(* Logix 5000 project; controller PLC_MCC1300_75F1 vendor 1 type 14 code 166 rev 32.11; software revision 32.04; part 77 of 83 *)
(* tags used below, declared in another part *)
   CM_AreaStackerToLine_JS1_Sync : CM_AreaStackerToLine;
   CM_ConveyorStackerToLine_JS1_Sync : CM_ConveyorStackerToLine;
   CONST_tPlant : UDT_PLANT_CONSTANTS;
   GP_AccessArea_M311S : GP_AccessArea;
   GP_AccessArea_M311S_STC : GP_AccessArea_STC;
   GP_AccessArea_M316S : GP_AccessArea;
   GP_AccessArea_M316S_STC : GP_AccessArea_STC;
   GP_OB_InitializeMain : GP_OB_Initialize;
   GP_TrackingGetLength : GP_TrackingGetLength;
   M302SpeedUp : MAC_SpeedUp;
   M30xTrimDeck : MAC_TrimmingDeck[5];
   M310B : MAC_Conveyor;
   M310B_ALM : MAC_Conveyor_ALM;
   M310B_HMW : MAC_Conveyor_HMW;
   M310Popup : MAC_Popup_ZC[2];
   M311 : MAC_Conveyor;
   M311_ALM : MAC_Conveyor_ALM;
   M311_HMW : MAC_Conveyor_HMW;
   M311A : MAC_Rotator;
   M311A_ALM : MAC_Rotator_ALM;
   M312 : MAC_Conveyor_Single;
   M312_ALM : MAC_Conveyor_ALM;
   M312_HMW : MAC_Conveyor_HMW;
   M316 : MAC_Conveyor;
   M316A : MAC_Rotator;
   M317 : MAC_Conveyor_Single;
   xAlwaysON : BOOL;
   Z300_Conveyor : UDT_StandConv[29];
   Z300_Conveyor_ALM : MAC_Conveyor_ZC_ALM[29];
   Z300_Conveyor_HMW : MAC_Conveyor_ZC_HMW[29];
   Z300_LineTracking : UDT_LINE_TRACKING;
   Z301 : MAC_Zone_ML;
   Z301_HMR : MAC_Zone_ML_HMR;
   Z301_HMW : MAC_Zone_ML_HMW;
   Z311S : MAC_SafetyAccess;
   Z311S_ALM : MAC_SafetyAccess_ALM;
   Z311S_HMR : MAC_SafetyAccess_HMR;
   Z311S_INPUT_xAccessReqRotator : BOOL;
   Z311S_INPUT_xSafetyAreaRotator : BOOL;
   Z311S_OUTPUT_xEL_AccessAcceptedRotator : BOOL;
   Z311S_OUTPUT_xHL_AccessAcceptedRotator : BOOL;
   Z311S_OUTPUT_xHL_SafetyAreaRotatorNOK : BOOL;
   Z316S : MAC_SafetyAccess;
   Z316S_ALM : MAC_SafetyAccess_ALM;
   Z316S_HMR : MAC_SafetyAccess_HMR;
   Z316S_INPUT_xAccessReqRotator : BOOL;
   Z316S_INPUT_xSafetyAreaRotator : BOOL;
   Z316S_OUTPUT_xEL_AccessAcceptedRotator : BOOL;
   Z316S_OUTPUT_xHL_AccessAcceptedRotator : BOOL;
   Z316S_OUTPUT_xHL_SafetyAreaRotatorNOK : BOOL;
   Z401 : MAC_Zone;
   Z401_ALM : MAC_Zone_ALM;
   Z401_HMR : MAC_Zone_HMR;
   Z401_HMW : MAC_Zone_HMW;
   Z401_INPUT_xMainLineEmergencyON : BOOL;
   Z401_OUTPUT_xMCC_SafetyPanel1 : BOOL;
   Z402 : MAC_Zone;
(* MainProgram, continued *)

   54: XIC(Z300_Conveyor_HMW[7].xLocalCleaningRequest)XIC(Z300_Conveyor[0].tIN_Zone.xCleanZoneAccepted)OTE(Z300_Conveyor_HMW[8].xLocalCleaningRequest);
   // M312 Cleaning Enabled
   55: XIC(Z300_Conveyor_HMW[8].xLocalCleaningRequest)XIC(Z300_Conveyor[0].tIN_Zone.xCleanZoneAccepted)[OTE(Z300_Conveyor_HMW[9].xLocalCleaningRequest) ,OTE(Z300_Conveyor_HMW[10].xLocalCleaningRequest) ];
   56: XIC(Z300_Conveyor_HMW[10].xLocalCleaningRequest)XIC(Z300_Conveyor[0].tIN_Zone.xCleanZoneAccepted)OTE(Z300_Conveyor_HMW[11].xLocalCleaningRequest);
   57: XIC(Z301.ST_xReqCleaning)XIC(Z300_Conveyor[0].ST_xCleaningConditionOK)XIC(Z300_Conveyor[1].ST_xCleaningConditionOK)XIC(Z300_Conveyor[2].ST_xCleaningConditionOK)XIC(Z300_Conveyor[3].ST_xCleaningConditionOK)XIC(Z300_Conveyor[4].ST_xCleaningConditionOK)XIC(Z300_Conveyor[5].ST_xCleaningConditionOK)XIC(Z300_Conveyor[6].ST_xCleaningConditionOK)XIC(Z300_Conveyor[7].ST_xCleaningConditionOK)XIC(Z300_Conveyor[8].ST_xCleaningConditionOK)XIC(Z300_Conveyor[9].ST_xCleaningConditionOK)XIC(Z300_Conveyor[10].ST_xCleaningConditionOK)XIC(Z300_Conveyor[11].ST_xCleaningConditionOK)XIC(M30xTrimDeck[0].ST_xCleaningConditionOK)XIC(M30xTrimDeck[1].ST_xCleaningConditionOK)XIC(M30xTrimDeck[2].ST_xCleaningConditionOK)XIC(M30xTrimDeck[3].ST_xCleaningConditionOK)XIC(M30xTrimDeck[4].ST_xCleaningConditionOK)OTE(Z301.ST_xCleaningConditionOK);
   58: XIC(Z301.ST_xReqCleaning)XIC(Z301.ST_xCleaningConditionOK)[OTL(Z301.ST_xCleaningAccepted) ,OTL(M302SpeedUp.ST_xFirstGlassAfterClean) ,OTE(Z301.OS_xCleaningAccepted) ];
   59: XIC(Z301.ST_xReqCleaning)XIC(Z301.ST_xCleaningAccepted)GP_TrackingGetLength(GP_TrackingGetLength,Z300_LineTracking,0,11)JSR(sbrTrackingPlateCleaning,4,0,GP_TrackingGetLength.OUT_dLength_cmm,0,0);
   // #####_HMI_STATUSES_#####
   60: NOP();
   61: XIC(Z301.ST_xZoneError)OTE(Z301_HMR.xZoneAlarm);
   62: XIC(Z301.ST_xCleaningAccepted)OTE(Z301_HMR.xCleaningEnabled);
   63: [MOV(0,Z301_HMR.dCabinetState) ,[XIC(Z300_Conveyor_ALM[0].rgxStoppingFault_M[0].x1) ,XIC(Z300_Conveyor_ALM[1].rgxStoppingFault_M[0].x1) ,XIC(Z300_Conveyor_ALM[2].rgxStoppingFault_M[0].x1) ,XIC(Z300_Conveyor_ALM[3].rgxStoppingFault_M[0].x1) ,XIC(Z300_Conveyor_ALM[4].rgxStoppingFault_M[0].x1) ,XIC(Z300_Conveyor_ALM[5].rgxStoppingFault_M[0].x1) ,XIC(Z300_Conveyor_ALM[5].rgxStoppingFault_M[1].x1) ,XIC(Z300_Conveyor_ALM[6].rgxStoppingFault_M[0].x1) ,XIC(Z300_Conveyor_ALM[7].rgxStoppingFault_M[0].x1) ,XIC(Z300_Conveyor_ALM[8].rgxStoppingFault_M[0].x1) ,XIC(Z300_Conveyor_ALM[9].rgxStoppingFault_M[0].x1) ,XIC(Z300_Conveyor_ALM[10].rgxStoppingFault_M[0].x1) ,XIC(Z300_Conveyor_ALM[11].rgxStoppingFault_M[0].x1) ,XIC(Z300_Conveyor_ALM[11].rgxStoppingFault_M[1].x1) ] MOV(2,Z301_HMR.dCabinetState) ,XIC(Z301.OUTPUT_xMCCSafetyLamp) MOV(1,Z301_HMR.dCabinetState) ];
   64: [MOV(0,Z301_HMR.dZoneMode) ,XIC(Z301.ST_xManuModeAccepted) MOV(1,Z301_HMR.dZoneMode) ,XIC(Z301.ST_xAutoModeAccepted) MOV(4,Z301_HMR.dZoneMode) ,XIC(Z301.ST_xManuModeReq) MOV(8,Z301_HMR.dZoneMode) ];
   65: [XIC(Z301.ST_xCycleON) MOV(1,Z301_HMR.dZoneState) ,XIO(Z301.ST_xCycleON) MOV(2,Z301_HMR.dZoneState) ,XIC(Z301.ST_xStartCycleRequest) XIO(Z301.ST_xCycleON) MOV(4,Z301_HMR.dZoneState) ,XIC(Z301.ST_xStopCycleRequest) XIC(Z301.ST_xCycleON) MOV(8,Z301_HMR.dZoneState) ,XIO(Z301.INPUT_xMainEmergencyON) MOV(1024,Z301_HMR.dZoneState) ];
   66: [MOV(2,Z301_HMR.dCleaningState) ,XIC(Z301.ST_xCleaningAccepted) MOV(1,Z301_HMR.dCleaningState) ,XIC(Z301.ST_xReqCleaning) MOV(4,Z301_HMR.dCleaningState) ];
   67: [MOV(Z301_HMW.dManualSpeed_mm_min,Z301_HMR.dManualSpeed_mm_min) ,LES(Z301_HMR.dManualSpeed_mm_min,CONST_tPlant.dMinLehrSpeed_mm_min) MOV(CONST_tPlant.dMinLehrSpeed_mm_min,Z301_HMR.dManualSpeed_mm_min) ,GRT(Z301_HMR.dManualSpeed_mm_min,CONST_tPlant.dMaxLineSpeed_mm_min) MOV(CONST_tPlant.dMaxLineSpeed_mm_min,Z301_HMR.dManualSpeed_mm_min) ];
   68: XIC(Z301.ST_xManuModeAccepted)XIC(Z301_HMW.rgxMan.0)XIC(Z300_Conveyor[0].ST_xRotationFeedback)XIC(Z300_Conveyor[1].ST_xRotationFeedback)XIC(Z300_Conveyor[2].ST_xRotationFeedback)XIC(Z300_Conveyor[3].ST_xRotationFeedback)XIC(Z300_Conveyor[4].ST_xRotationFeedback)XIC(Z300_Conveyor[5].ST_xRotationFeedback)XIC(Z300_Conveyor[6].ST_xRotationFeedback)XIC(Z300_Conveyor[7].ST_xRotationFeedback)XIC(Z300_Conveyor[8].ST_xRotationFeedback)XIC(Z300_Conveyor[9].ST_xRotationFeedback)XIC(Z300_Conveyor[10].ST_xRotationFeedback)XIC(Z300_Conveyor[11].ST_xRotationFeedback)OTE(Z301_HMR.rgxMan.0);
END_ROUTINE

ROUTINE Z311S_Alarm   (* ladder *)
   0: XIC(Z401.tmON_ResetAlarm.DN)FLL(0,Z311S_ALM,1);
   1: XIC(Z401.ST_xEnableControlError)XIO(Z311S_INPUT_xSafetyAreaRotator)XIO(GP_AccessArea_M311S_STC.ST_xAccessAccepted)OTE(Z311S_ALM.rgxFault[0].1);
END_ROUTINE

ROUTINE Z311S_Logic   (* ladder *)
   // #####_ALARMS_#####
   0: NOP();
   1: JSR(Z311S_Alarm,0);
   // #####_PHASES_&_LOGICS_#####
   2: NOP();
   // M311S - Taglia solo rotatore e salita/discesa rotatore
   3: XIC(M311A.ST_xConditionOKStopCycle)XIC(M312.ST_xConditionOKStopCycle)OTE(Z311S.xMxx0S_ConditionOK);
   4: GP_AccessArea(GP_AccessArea_M311S,GP_AccessArea_M311S_STC,Z311S_INPUT_xAccessReqRotator,0,Z311S.xMxx0S_ConditionOK,0,GP_OB_InitializeMain.OUT_xClock_800ms,Z311S_OUTPUT_xHL_AccessAcceptedRotator);
   5: XIC(GP_AccessArea_M311S_STC.ST_xAccessAccepted)OTE(Z311S_OUTPUT_xEL_AccessAcceptedRotator);
   6: XIO(Z311S_INPUT_xSafetyAreaRotator)XIO(GP_AccessArea_M311S_STC.ST_xAccessRequest)XIO(GP_AccessArea_M311S_STC.ST_xAccessAccepted)OTE(Z311S_OUTPUT_xHL_SafetyAreaRotatorNOK);
   // M311S - taglia M312 (trasportatore verso stk) - M312 (salita/discesa) - M312 (sollevamento popup)
   7: XIC(M311.ST_xConditionOKStopCycle)XIC(M312.ST_xConditionOKStopCycle)OTE(Z311S.xMxx1S_ConditionOK);
   // #####_HMI_STATUS_#####
   8: NOP();
   9: [MOV(1,Z311S_HMR.iMxx0S_State) ,XIC(GP_AccessArea_M311S_STC.ST_xAccessRequest) MOV(2,Z311S_HMR.iMxx0S_State) ,XIC(GP_AccessArea_M311S_STC.ST_xAccessAccepted) MOV(8,Z311S_HMR.iMxx0S_State) ,XIO(Z311S_INPUT_xSafetyAreaRotator) MOV(4,Z311S_HMR.iMxx0S_State) ];
END_ROUTINE

ROUTINE Z316S_Alarm   (* ladder *)
   0: XIC(Z402.tmON_ResetAlarm.DN)FLL(0,Z316S_ALM,1);
   1: XIC(Z402.ST_xEnableControlError)XIO(Z316S_INPUT_xSafetyAreaRotator)XIO(GP_AccessArea_M316S_STC.ST_xAccessAccepted)OTE(Z316S_ALM.rgxFault[0].1);
END_ROUTINE

ROUTINE Z316S_Logic   (* ladder *)
   // #####_ALARMS_#####
   0: NOP();
   1: JSR(Z316S_Alarm,0);
   // #####_PHASES_&_LOGICS_#####
   2: NOP();
   // M316S - Taglia solo rotatore e salita/discesa rotatore
   3: XIC(M316A.ST_xConditionOKStopCycle)XIC(M317.ST_xConditionOKStopCycle)OTE(Z316S.xMxx0S_ConditionOK);
   4: GP_AccessArea(GP_AccessArea_M316S,GP_AccessArea_M316S_STC,Z316S_INPUT_xAccessReqRotator,0,Z316S.xMxx0S_ConditionOK,0,GP_OB_InitializeMain.OUT_xClock_800ms,Z316S_OUTPUT_xHL_AccessAcceptedRotator);
   5: XIC(GP_AccessArea_M316S_STC.ST_xAccessAccepted)OTE(Z316S_OUTPUT_xEL_AccessAcceptedRotator);
   6: XIO(Z316S_INPUT_xSafetyAreaRotator)XIO(GP_AccessArea_M316S_STC.ST_xAccessRequest)XIO(GP_AccessArea_M316S_STC.ST_xAccessAccepted)OTE(Z316S_OUTPUT_xHL_SafetyAreaRotatorNOK);
   // M311S - taglia M312 (trasportatore verso stk) - M312 (salita/discesa) - M312 (sollevamento popup)
   7: XIC(M316.ST_xConditionOKStopCycle)XIC(M317.ST_xConditionOKStopCycle)OTE(Z316S.xMxx1S_ConditionOK);
   // #####_HMI_STATUS_#####
   8: NOP();
   9: [MOV(1,Z316S_HMR.iMxx0S_State) ,XIC(GP_AccessArea_M316S_STC.ST_xAccessRequest) MOV(2,Z316S_HMR.iMxx0S_State) ,XIC(GP_AccessArea_M316S_STC.ST_xAccessAccepted) MOV(8,Z316S_HMR.iMxx0S_State) ,XIO(Z316S_INPUT_xSafetyAreaRotator) MOV(4,Z316S_HMR.iMxx0S_State) ];
END_ROUTINE

ROUTINE Z401_Alarm   (* ladder *)
   0: XIC(Z401.tmON_ResetAlarm.DN)FLL(0,Z401_ALM,1);
END_ROUTINE

ROUTINE Z401_Logic   (* ladder *)
   // #####_COSTANTS_#####
   0: NOP();
   // #####_MATCH_#####
   1: NOP();
   // #####_ALARMS_#####
   2: NOP();
   3: XIC(Z401_HMW.xResetErrorRequest)[OTU(Z401_HMW.xResetErrorRequest) ,TOF(Z401.tmON_ResetAlarm,?,?) ];
   4: XIC(Z401.tmON_24Vdc.DN)XIC(Z401.tmON_400Vca.DN)XIC(Z401.tmON_EmergencyOK.DN)OTE(Z401.ST_xEnableControlError);
   5: JSR(Z401_Alarm,0);
   // #####_HMI_LOGICS_#####
   6: NOP();
   // #####_STATUSES_#####
   7: NOP();
   8: [NEQ(Z401_ALM.rgxEmergency[0],0) ,NEQ(Z401_ALM.rgxFault[0],0) ,NEQ(Z401_ALM.rgxWarning[0],0) ,XIC(M310Popup[0].ST_xMachineAlarm) ,XIC(M310Popup[1].ST_xMachineAlarm) ,XIC(M311.ST_xMachineAlarm) ,XIC(M311A.ST_xMachineAlarm) ,XIC(M312.ST_xMachineAlarm) ]OTE(Z401.ST_xZoneError);
   // #####_ZONE MODALITY_#####
   9: NOP();
   // Selector manual mode
   10: XIC(Z401_HMW.xManualModeRequest)OTL(Z401.ST_xSelectionManualMode)OTU(Z401.ST_xSelectionAutomaticMode)OTU(Z401_HMW.xManualModeRequest);
   // Selector automatic mode
   11: XIC(Z401_HMW.xAutomaticModeRequest)OTL(Z401.ST_xSelectionAutomaticMode)OTU(Z401.ST_xSelectionManualMode)OTU(Z401_HMW.xAutomaticModeRequest);
   // Condition Ok for manual mode
   12: [XIC(Z401.ST_xConditionOKStopCycle) ,XIO(Z401.ST_xCycleON) ]OTE(Z401.ST_xConditionOkManualMode);
   // Manual mode accepted
   13: XIC(Z401.ST_xSelectionManualMode)[XIO(Z401.ST_xManualModeAccepted) OTE(Z401.ST_xManualModeRequest) ,[XIC(Z401.ST_xConditionOkManualMode) ,XIC(Z401.ST_xManualModeAccepted) ] OTE(Z401.ST_xManualModeAccepted) ];
   // Auto mode accepted
   14: XIO(Z401.ST_xManualModeAccepted)[XIC(Z401.ST_xSelectionAutomaticMode) ,XIC(Z401.ST_xAutoModeAccepted) ][OTE(Z401.ST_xAutoModeAccepted) ,ONS(Z401.OSR_xAutomaticMode) OTE(Z401.OS_xAutomaticMode) ];
   // Set all manual command for iFix
   15: XIC(Z401.ST_xManualModeAccepted)OTL(M310B_HMW.xEnableDisableManualCommand)OTL(M311_HMW.xEnableDisableManualCommand)OTL(M312_HMW.xEnableDisableManualCommand);
   // Reset all manual command for iFix
   16: XIC(Z401.OS_xAutomaticMode)OTU(M310B_HMW.xEnableDisableManualCommand)OTU(M311_HMW.xEnableDisableManualCommand)OTU(M312_HMW.xEnableDisableManualCommand);
   // #####_LOGICS_#####
   17: NOP();
   18: [XIC(Z401_HMW.xStartCycleRequest) ,XIC(CM_AreaStackerToLine_JS1_Sync.xSB_LineCycle) ]OTE(Z401.OS_xStartCycle);
   19: [XIC(Z401_HMW.xStopCycleRequest) ,XIC(CM_AreaStackerToLine_JS1_Sync.xSB_StopLineCycle) ]OTE(Z401.OS_xStopCycle);
   20: [XIC(Z401.tmON_ForceStop.DN) ONS(Z401.OSR_xForceStopCycle) ,XIC(Z401_HMW.xForceStopCycle) ]OTE(Z401.OS_xForceStopCycle);
   21: XIO(Z401.OS_xForceStopCycle)XIC(Z401.tmON_24Vdc.DN)XIC(Z401.tmON_400Vca.DN)XIC(Z401.tmON_EmergencyOK.DN)OTE(Z401.ST_xConditionOkCycleON);
   22: [XIC(Z401.OS_xStartCycle) ,XIC(Z401.ST_xStartCycleRequest) ]XIC(Z401.ST_xConditionOkCycleON)XIO(Z401.ST_xCycleON)XIO(Z401.OS_xStopCycle)OTE(Z401.ST_xStartCycleRequest);
   23: [XIC(Z401.OS_xStopCycle) ,XIC(Z401.ST_xStopCycleRequest) ]XIC(Z401.ST_xCycleON)XIO(Z401.ST_xStartCycleRequest)OTE(Z401.ST_xStopCycleRequest);
   24: XIC(M310B.ST_xConditionOKStopCycle)XIC(M311.ST_xConditionOKStopCycle)XIC(M311A.ST_xConditionOKStopCycle)XIC(M312.ST_xConditionOKStopCycle)XIC(CM_ConveyorStackerToLine_JS1_Sync.xConditionOkForStopCycle)OTE(Z401.ST_xConditionOKStopCycle);
   25: [XIC(Z401.ST_xStopCycleRequest) XIC(Z401.ST_xConditionOKStopCycle) ,XIC(Z401_HMW.xForceStopCycle) ]OTE(Z401.ST_xStopCycleAccepted);
   // Reimpostare tempo a 15 secondi
   26: [XIC(Z401.ST_xStartCycleRequest) ,XIC(Z401.ST_xCycleON) ]XIC(Z401.ST_xConditionOkCycleON)XIO(Z401.ST_xStopCycleAccepted)XIO(Z401.ST_xManualModeAccepted)[TON(Z401.tmON_Cycle,?,?) ,XIC(Z401.tmON_Cycle.DN) OTE(Z401.ST_xCycleON) ];
   27: XIC(Z401.ST_xCycleON)XIO(Z401.ST_xManualModeRequest)XIO(Z401.ST_xStopCycleRequest)OTE(Z401.ST_xConditionOkPhaseAdvancement);
   28: XIC(Z401.ST_xCycleON)[XIC(M310B.ST_xCleaningAccepted) ,XIO(M310B.ST_xReqCleaning) ][XIC(M311.ST_xCleaningAccepted) ,XIO(M311.ST_xReqCleaning) ][XIC(M312.ST_xCleaningAccepted) ,XIO(M312.ST_xReqCleaning) ]OTE(Z401.ST_xCleaningConditionOK);
   // Speed manager
   29: [MOV(Z401_HMW.dLineSpeed_mm_min,Z401_HMR.dLineSpeed_mm_min) ,LES(Z401_HMR.dLineSpeed_mm_min,35000) MOV(35000,Z401_HMR.dLineSpeed_mm_min) ,GRT(Z401_HMR.dLineSpeed_mm_min,60000) MOV(60000,Z401_HMR.dLineSpeed_mm_min) ];
   // #####_CLEANING_#####
   30: NOP();
   31: XIO(Z401.ST_xCleaningAccepted)XIC(Z401_HMW.xStartCleanZoneRequest)[MOV(Z401_HMW.dCleaningSelection,Z401_HMR.dCleaningSelection) ,OTL(Z401.ST_xReqCleaning) ];
   32: XIC(Z401.ST_xReqCleaning)XIC(Z401.ST_xCleaningConditionOK)[OTL(Z401.ST_xCleaningAccepted) ,OTU(Z401.ST_xReqCleaning) ,OTL(M310B_HMW.xLocalCleaningRequest) ,OTL(M311_HMW.xLocalCleaningRequest) ,OTL(M312_HMW.xLocalCleaningRequest) ];
   33: XIC(Z401_HMW.xStopCleanZoneRequest)[OTU(Z401.ST_xReqCleaning) ,OTU(Z401.ST_xCleaningAccepted) ,MOV(0,Z401_HMW.dCleaningSelection) ,OTU(M310B_HMW.xLocalCleaningRequest) ,OTU(M311_HMW.xLocalCleaningRequest) ,OTU(M311_HMW.xLocalCleaningRequest) ];
   34: XIC(xAlwaysON)[OTU(Z401_HMW.xStartCycleRequest) ,OTU(Z401_HMW.xStopCycleRequest) ,OTU(Z401_HMW.xStartCleanZoneRequest) ,OTU(Z401_HMW.xForceStopCycle) ,OTU(Z401_HMW.xStopCleanZoneRequest) ];
   // #####_HMI_STATUSES_#####
   35: NOP();
   36: XIC(Z401.ST_xZoneError)OTE(Z401_HMR.xZoneAlarm);
   37: [XIC(Z401.ST_xCleaningAccepted) ,XIC(M310B.ST_xCleaningAccepted) XIC(M311.ST_xCleaningAccepted) XIC(M312.ST_xCleaningAccepted) ]OTE(Z401_HMR.xCleaningEnabled);
   38: [MOV(0,Z401_HMR.dCabinetState1) ,[XIC(M310B_ALM.rgxStoppingFault_M[0].1) ,XIC(M311_ALM.rgxStoppingFault_M[0].1) ,XIC(M311A_ALM.rgxStoppingFault_M[0].1) ,XIC(M312_ALM.rgxStoppingFault_M[0].1) ] MOV(2,Z401_HMR.dCabinetState1) ,XIC(Z401_OUTPUT_xMCC_SafetyPanel1) MOV(1,Z401_HMR.dCabinetState1) ];
   39: [XIC(Z401.ST_xManualModeAccepted) MOV(1,Z401_HMR.dZoneMode) ,XIC(Z401.ST_xAutoModeAccepted) MOV(4,Z401_HMR.dZoneMode) ,XIC(Z401.ST_xManualModeRequest) MOV(8,Z401_HMR.dZoneMode) ];
   40: [MOV(2,Z401_HMR.dZoneState) ,XIC(Z401.ST_xStartCycleRequest) XIO(Z401.ST_xCycleON) MOV(4,Z401_HMR.dZoneState) ,XIC(Z401.ST_xCycleON) MOV(1,Z401_HMR.dZoneState) ,XIC(Z401.ST_xStopCycleRequest) MOV(8,Z401_HMR.dZoneState) ,XIO(Z401_INPUT_xMainLineEmergencyON) MOV(1024,Z401_HMR.dZoneState) ];
   41: [[XIC(Z401.ST_xCleaningAccepted) ,XIC(M310B.ST_xCleaningAccepted) XIC(M311.ST_xCleaningAccepted) XIC(M312.ST_xCleaningAccepted) ] MOV(1,Z401_HMR.dCleaningState) ,XIO(Z401.ST_xCleaningAccepted) MOV(2,Z401_HMR.dCleaningState) ,XIC(Z401.ST_xReqCleaning) XIO(Z401.ST_xCleaningAccepted) MOV(4,Z401_HMR.dCleaningState) ];
